// TIA Portal project "S7_1516_LECTOR620_DI" (V15) (continued)
VERSION : 1.2
// The function block use a Profinet/Probibus connection to communicate with a SICK AutoIdent
// device. The FB makes it possible to send and receive sensor data. The Confirmed Messaging 
// protocol (CM-Protocol) is used to receive even long fragmented read results.
// The function block use a Profinet/Probibus connection to communicate with a SICK AutoIdent
// device. The FB makes it possible to send and receive sensor data.
   VAR_INPUT
      HWInputIdent : Hw_Io;   // Hardware identification number of the input module
      HWInputLength : USInt;   // Size of the input module
      HWOutputIdent : Hw_Io;   // Hardware identification number of the output module
      HWOutputLength : USInt;   // Size of the output module
      TOut : Time := T#5s;   // Time out
      Req : Bool;   // A positive edge starts the request
      CommandLength : UInt;   // Byte length of the command / Command length in byte
   END_VAR
   VAR_OUTPUT
      RdDone : Bool;   // Reading result arrived / Positive edge: A reading result sent by the device was received
      RdLength : Int;   // Byte length of the reading result / Length of the reading result in byte
      ReqDone : Bool;   // Requested data available / Indicates whether a CoLa command was sent and an answer was received
      ReqBusy : Bool;   // Request busy / Request processing
      ReqLength : Int;   // Byte length of the requested data / Length of an answer telegram in byte
      Error : Bool;   // Error / Error detected
      Errorcode : DWord;   // Error code / Error code (see documentation)
   END_VAR
   VAR_IN_OUT
      arrCommand : Array[0..499] of Byte;   // Contain the transmitted CoLa command without STX/ETX framing
      arrRecord : Array[0..499] of Byte;   // Contain the received telegram
   END_VAR
   VAR
      bTriggerReq : Bool := false;   // Rising edge detection
      bTriggerReqMem : Bool := false;   // Rising edge detection
      bReadFrag : Bool;   // Fragmentation is needed (Read)
      bWriteFrag : Bool;   // Fragmentation is needed (Write)
      bReqBusyMem : Bool;
      iReadStep : USInt;   // Current step (Read)
      iWriteStep : USInt;   // Current step (Write)
      iReadIndex : UInt;   // Index (Read)
      iWriteIndex : UInt;   // Index (Write)
      iReadHeaderLength : UInt;   // Header length of the CM-Protocol (Read)
      iWriteHeaderLength : UInt;   // Header length of the CM-Protocol (Write)
      iReadFragmentLength : UInt;   // Length of the current fragment (Read)
      iWriteFragmentLength : UInt;   // Length of the current fragment (Write)
      iRecordSize : UInt;   // Length of the record array
      iCommandSize : UInt;   // Length of the command array
      nTempErrorCode : DWord;   // Temporarily error code
      arrInputImage : Array[0..127] of Byte;   // Process data input image
      arrOutputImage : Array[0..127] of Byte;   // Process data output image
      fbTimeout : TON_TIME;   // Instance: Timer on delay (Time out)
   END_VAR
   VAR_TEMP
      iTemp1 : Int;   // Temporarily variable
      iTemp2 : UDInt;   // Temporarily variable
      iTemp3 : UDInt;   // Temporarily variable
   END_VAR
BEGIN
   (*===========================================================================================
   Name:   SICK_CCOMM_PNDP
   Author: SICK AG
   =============================================================================================
   Description: 
   The function block use a Profinet/Probibus connection to communicate with a SICK AutoIdent
   device. The FB makes it possible to send and receive sensor data. The Confirmed Messaging 
   protocol (CM-Protocol) is used to receive even long fragmented read results.

   Send a command:
   The "Req" parameter must be triggered with a rising edge (signal change FALSE to TRUE) in 
   order to carry out the function. For the time during which a valid response has yet to be 
   received from the device, the "ReqBusy" parameter is used to signal  that a response is still 
   pending. The module signals the "ReqDone" = TRUE output parameter when the function has been 
   successfully completed. If data was requested by the device, this data is copied into the 
   Record (arrRecord). The "ReqDone" indicates that new data has been received  for a PLC cycle.
   Only one CoLa-A command request can be send to the same device at one time. 

   Receive a reading result:
   Data sent via trigger command or directly by the device (e.g., direct trigger via a light 
   barrier) is stored in the Record (arrRecord). The "RdDone" output indicates that new data 
   has been received for a PLC cycle. The data sent by the device can be changed or adapted in 
   output format of SOPAS-ET. 

   This AOI supports the folowing SICK devices:
   - Lector6xx
   - RFU6xx
   - CLV6xx 
   - RFH6xx
   =============================================================================================
   Confirmed Messaging Protocol definitions:
   arrInputImage[0]        = Status byte 
   arrInputImage[1]        = Receive counter
   arrInputImage[2]        = Transmit counter back
   arrInputImage[3]        = Command length LSB
   arrInputImage[4]        = Command length MSB
   arrInputImage[5..127]   = Device response (CoLa-A)

   arrOutputImage[0]       = Status byte 
   arrOutputImage[1]       = Receive counter back
   arrOutputImage[2]       = Transmit counter
   arrOutputImage[3]       = Command length LSB
   arrOutputImage[4]       = Command length MSB
   arrOutputImage[5..127]  = Device request (CoLa-A)
   =============================================================================================
   Version history:
   Date       | Version | Created under               | Author  | Remark
   ---------------------------------------------------------------------------------------------
   16/01/2014 | V1.0    | TIA Portal V12 SP1 Update 2 | SICK AG | Initial version
   07/08/2014 | V1.1    | TIA Portal V12 SP1 Update 4 | SICK AG | Replace R_TRIG function 
   22/04/2015 | V1.2    | TIA Portal V12 SP1 Update 4 | SICK AG | Avoid warnings that occur with 
                                                                  TIA V13
   ============================================================================================*)

   (*===================================== INITIALISATION =====================================*)
   #iRecordSize:= 500;   (*Length of the arrRecord array*)
   #iCommandSize:= 500;  (*Length of the arrCommand array*)

   #RdDone:= false;
   #iReadStep:= 0;

   (*Rising edge detection of the request flag*)
   #bTriggerReq:= #Req AND NOT #bTriggerReqMem;
   #bTriggerReqMem:= #Req;

   (*Error detection*)
   IF #nTempErrorCode <>16#0000_0000 THEN
     #ReqDone:= false;
     #ReqBusy:= false;
     #bReqBusyMem:= false;
     #Error:= true;
     #Errorcode:= #nTempErrorCode;
     #nTempErrorCode:= 16#0000_0000;
     #ReqLength:= 0;
     #iWriteStep:= 0;
     RETURN;
   END_IF;

   (*Time out detection*)
   #fbTimeout(IN:=#bReqBusyMem, PT:=#TOut);
   IF #fbTimeout.Q THEN
     #nTempErrorCode:= 16#0000_0001; (*Error: Time out*) 
   END_IF;

   (*Check the hardware ident length of the input module*)
   IF #HWInputLength <8 OR #HWInputLength >128 THEN
     #nTempErrorCode:= 16#0000_0002; (*Error: Incorrect module input length*)
   END_IF;

   (*Check the hardware ident length of the output module*)
   IF #HWOutputLength <8 OR #HWOutputLength >128 THEN
     #nTempErrorCode:= 16#0000_0003; (*Error: Incorrect module output length*)
   END_IF;

   (*Error detected*)
   IF #nTempErrorCode <>16#0000_0000 THEN
     RETURN;
   END_IF;


   (*===================================== COMMUNICATION ======================================*)
   (*Set output data*)
   #iTemp1:= DPWR_DAT(LADDR:= #HWOutputIdent, RECORD:= #arrOutputImage);
   IF #iTemp1 <>0 THEN
     #nTempErrorCode.%W1:= #iTemp1;
     #nTempErrorCode.%W0:= 16#0004; (*Error: Set output data via DPWR_DAT*)
     RETURN;
   END_IF;

   (*Get input data*)
   #iTemp1:= DPRD_DAT(LADDR:= #HWInputIdent, RECORD=> #arrInputImage);
   IF #iTemp1 <>0 THEN
     #nTempErrorCode.%W1:= #iTemp1;
     #nTempErrorCode.%W0:= 16#0005; (*Error: Get input data via DPRD_DAT*)
     RETURN;
   END_IF;

   (*Receive counter ==0 && Receive counter back <>0*)
   IF #arrInputImage[1] =0 AND #arrOutputImage[1] <>0 THEN
     #arrOutputImage[1]:= #arrInputImage[1]; (*Recive counter => Receive counter back*)
     RETURN;
   END_IF;

   (*Transmit counter <> Transmit counter back*)
   IF NOT #bReqBusyMem AND (#arrInputImage[2] <> #arrOutputImage[2]) THEN
     #arrOutputImage[2]:= 0; (*0 => Transmit counter*)
     RETURN;
   END_IF;


   (*============================== HANDLING OF THE RECEIVED DATA =============================*)
   (*New telegram available*)
   IF NOT (#arrInputImage[1] = #arrOutputImage[1]) THEN

     (*Reset error every incoming telegram (Read only mode, e.g. for hand held scanners)*)
     IF #CommandLength <=0 THEN
       #Error:= false;
       #Errorcode:= 16#0000_0000;
     END_IF;

     (*Confirm the receive counter*)
     #arrOutputImage[1]:= #arrInputImage[1];

     (*Get telegram length from the received header*)
     #iReadHeaderLength.%B0:= #arrInputImage[3];
     #iReadHeaderLength.%B1:= #arrInputImage[4];

     (*Check if fragmentation is not active at the moment*)
     IF NOT #bReadFrag THEN
       #iReadIndex:= 0;

       (*Check if fragmentation is needed*)
       IF (#HWInputLength-5) < #iReadHeaderLength THEN
         #bReadFrag:= true;
       END_IF;
     END_IF;

     (*Fragmentation is needed*)
     IF #bReadFrag THEN
       IF (#HWInputLength-5) < #iReadHeaderLength THEN
         #iReadFragmentLength:= #HWInputLength-5;
       ELSE
         #iReadFragmentLength:= #iReadHeaderLength;
       END_IF;

     (*No fragmentation needed*)
     ELSE
       #iReadFragmentLength:= #iReadHeaderLength;
     END_IF;

     (*Copy input data into the output record*)
     IF (#iReadIndex+#iReadFragmentLength) <= #iRecordSize THEN
       MOVE_BLK(IN:= #arrInputImage[5], COUNT:= #iReadFragmentLength, OUT=> #arrRecord[#iReadIndex]);
     END_IF;

     (*Check if all data has been received*)
     IF (#HWInputLength-5) < #iReadHeaderLength THEN
       #iReadIndex:= #iReadIndex+#iReadFragmentLength;

     (*All data has been received*)
     ELSE
       #bReadFrag:= false;
       #iReadStep:= 1;
     END_IF;

     (*Incoming data filter*)
     (* - Check if the receiving telegram os a CoLa answer on a requested 
          comand or a reading result.

         sRA  sWA  sMA  sAN  sAI  sEA  sPX  s{   sSI  sSN  sFA
     sRN  X                                       X    X    X
     sRI  X                                       X    X    X
     sWN       X                                  X    X    X
     sWI       X                                  X    X    X
     sMN            X    X                        X    X    X
     sMI            X         X                   X    X    X
     sEN                           X              X    X    X
     sEI                           X              X    X    X
     sPE                                X         X    X    X
     s{                                      X    X    X    X
     *)
     IF #iReadStep =1 THEN
       (*Filter is only active, while requested data expected*)
       IF #bReqBusyMem THEN
         IF #CommandLength >3 THEN
           (*Get the prefix from the requested command (e.g. 'sRN '*)   
           #iTemp2.%B3:= #arrCommand[0];
           #iTemp2.%B2:= #arrCommand[1];
           #iTemp2.%B1:= #arrCommand[2];
           #iTemp2.%B0:= 16#20;

           (*Get the prefix from the command response (e.g. 'sRA ')*)
           #iTemp3.%B3:= #arrRecord[0];
           #iTemp3.%B2:= #arrRecord[1];
           #iTemp3.%B1:= #arrRecord[2];
           #iTemp3.%B0:= 16#20;
         ELSE
           #iTemp2:= 16#0000_0000;
           #iTemp3:= 16#0000_0000;
         END_IF;

         CASE #iTemp3 OF
         (*'s{  '*)
         16#737B2020:  IF #iTemp2 = 16#737B2020 THEN
                         #iReadStep:= 2; (*Command response*)
                       ELSE
                         #iReadStep:= 3; (*Reading result*)
                       END_IF;

         (*'sRA '*)
         16#73524120:  IF (#iTemp2 = 16#73524E20) OR (#iTemp2 = 16#73524920) THEN
                         #iReadStep:= 2; (*Command response*)
                       ELSE
                         #iReadStep:= 3; (*Reading result*)
                       END_IF;

         (*'sWA '*)
         16#73574120:  IF (#iTemp2 = 16#73574E20) OR (#iTemp2 = 16#73574920) THEN
                         #iReadStep:= 2; (*Command response*)
                       ELSE
                         #iReadStep:= 3; (*Reading result*)
                       END_IF;

         (*'sMA '*)
         16#734D4120:  IF (#iTemp2 = 16#734D4E20) OR (#iTemp2 = 16#734D4920) THEN
                         #iReadStep:= 2; (*Command response*)
                       ELSE
                         #iReadStep:= 3; (*Reading result*)
                       END_IF;

         (*'sAN '*)
         16#73414E20:  IF #iTemp2 = 16#734D4E20 THEN
                         #iReadStep:= 2; (*Command response*)
                       ELSE
                         #iReadStep:= 3; (*Reading result*)
                       END_IF;

         (*'sAI '*)
         16#73414920:  IF #iTemp2 = 16#734D4920 THEN
                         #iReadStep:= 2; (*Command response*)
                       ELSE
                         #iReadStep:= 3; (*Reading result*)
                       END_IF;

         (*'sEA '*)
         16#73454120:  IF (#iTemp2 = 16#73454E20) OR (#iTemp2 = 16#73454920) THEN
                         #iReadStep:= 2; (*Command response*)
                       ELSE
                         #iReadStep:= 3; (*Reading result*)
                       END_IF;

         (*'sPX '*)
         16#73505820:  IF #iTemp2 = 16#73504520 THEN
                         #iReadStep:= 2; (*Command response*)
                       ELSE
                         #iReadStep:= 3; (*Reading result*)
                       END_IF;

         (*'sSI '*)
         16#73534920:  #iReadStep:= 3; (*Reading result*)

         (*'sSN '*)
         16#73534E20:  #iReadStep:= 3; (*Reading result*)

         (*'sFA '*)
         16#73464120:  #iReadStep:= 2; (*Command response*)

         (*Invalid CoLa-A answer*)
         ELSE
           (*Check if a user defined command is used (Request == Response)*)
           FOR #iTemp1:= 0 TO UINT_TO_INT(#CommandLength-1) DO
             IF #arrCommand[#iTemp1] = #arrRecord[#iTemp1] THEN
               #iReadStep:= 2; (*Command response*)
             ELSE
               #iReadStep:= 3; (*Reading result*)
               EXIT;
             END_IF;
           END_FOR;
         END_CASE;

       (*Reading result*)
       ELSE
         #iReadStep:= 3;  (*Reading result*)
       END_IF;
     END_IF;

     (*Incoming telegram is a command response*)
     IF #iReadStep =2 THEN
       IF (#iReadIndex+#iReadFragmentLength) <= #iRecordSize THEN
         #ReqLength:= UDINT_TO_INT(#iReadIndex+#iReadFragmentLength);
         #ReqDone:= true;
         #ReqBusy:= false;
         #bReqBusyMem:= false;
       ELSE
         #nTempErrorCode:= 16#0000_0006; (*Error: Incoming command response > Record size*)
       END_IF;
     END_IF;

     (*Incoming telegram is a reading result*)
     IF #iReadStep =3 THEN
       IF (#iReadIndex+#iReadFragmentLength) <= #iRecordSize THEN
         #RdLength:= UDINT_TO_INT(#iReadIndex+#iReadFragmentLength);
         #RdDone:= true;
       ELSE
         #RdLength:= -1;
         #RdDone:= false;    
       END_IF;
     END_IF;
   END_IF;


   (*=========================== HANDLING OF THE DATA TO BE WRITTEN ===========================*)
   IF #bTriggerReq AND NOT #bReqBusyMem THEN
     #ReqDone:= false;
     #ReqBusy:= true;
     #bReqBusyMem:= true;
     #Error:= false;
     #Errorcode:= 16#0000_0000;
     #iWriteIndex:= 0;

     (*Check command length*)
     IF #CommandLength <=0 THEN
       #nTempErrorCode:= 16#0000_0007; (*Error: Command length <= 0*)
       RETURN;
     ELSIF #CommandLength > #iCommandSize THEN
       #nTempErrorCode:= 16#0000_0008; (*Error: Command length > command array*)
       RETURN;
     END_IF;

     (*Check if the the command telegram must be fragmented*)
     IF (#HWOutputLength-5) < #CommandLength THEN
       #iWriteFragmentLength:= #HWOutputLength-5;
     ELSE
       #iWriteFragmentLength:= #CommandLength;
     END_IF;

     #iWriteHeaderLength:= #CommandLength;
     #iWriteStep:= 1;  
   END_IF;

   (*Write step 1: Command transfer*)
   IF (#iWriteStep =1) AND(#arrInputImage[2] = #arrOutputImage[2]) THEN

     (*Copy command data into the output record*)
     IF((#iWriteIndex+#iWriteFragmentLength) <= #iCommandSize) AND (#iWriteFragmentLength <= (#HWOutputLength-5)) THEN
       MOVE_BLK(IN:= #arrCommand[#iWriteIndex], COUNT:= #iWriteFragmentLength, OUT=> #arrOutputImage[5]);
       (*Increment transmit counter*)
       IF #arrOutputImage[2] = 16#FF THEN
         #arrOutputImage[2]:= 16#01; (*Counter overflow, zero is skipped*)
       ELSE
         #arrOutputImage[2]:= #arrOutputImage[2]+1;
       END_IF;

       (*Set command/fragment length*)
       #arrOutputImage[3]:= #iWriteHeaderLength.%B0;
       #arrOutputImage[4]:= #iWriteHeaderLength.%B1;

       (*Next step*)
       #iWriteStep:= 2;
     ELSE
       #nTempErrorCode:= 16#0000_0009; (*Error: Fragmentation error*)
     END_IF;
       RETURN;
   END_IF;

   (*Write step 2: Fragmentation handling*)
   IF #iWriteStep =2 THEN

     (*Fragmentation is needed*)
     IF (#HWOutputLength-5) < #iWriteHeaderLength THEN
       #bWriteFrag:= true;

       (*Next index*)
       #iWriteIndex:= #iWriteIndex+#iWriteFragmentLength;

       (*Set next header length*)
       #iWriteHeaderLength:= #iWriteHeaderLength-#iWriteFragmentLength;

       (*Set next fragment length*)
       IF (#HWOutputLength-5) < #iWriteHeaderLength THEN
         #iWriteFragmentLength:= #HWOutputLength-5;
       ELSE
         #iWriteFragmentLength:= #iWriteHeaderLength;
       END_IF;

     (*Fragmentation is not needed*)
     ELSE
       #bWriteFrag:= false;
     END_IF;

     (*Next step*)
     #iWriteStep:= 3;
   END_IF;

   (*Write step 3: Check if the transmission of the command/fragment is done*)
   IF #iWriteStep =3 THEN

     (*Transmit counter back == Transmit counter*)
     IF #arrInputImage[2] = #arrOutputImage[2] THEN
       IF #bWriteFrag THEN
         #iWriteStep:= 1;
       ELSE
         #iWriteStep:= 0;
       END_IF;
     END_IF;
   END_IF;
END_FUNCTION_BLOCK

FUNCTION "SICK_GetValue" : Void   // FC10, SCL
TITLE = Get value
{ S7_Optimized_Access := 'TRUE' }
AUTHOR : SICKAG
FAMILY : Ident
VERSION : 1.0
// This function is needs to get a value out of a SICK CoLa command.
   VAR_INPUT
      iTelegramLength : UInt;   // Length of the source telegram
      iValueLength : USInt;   // ASCII length of the value [1..8] = Fix length | [0]= Variable
      arrData : Array[0..499] of Byte;   // Data record (contains the whole CoLa telegram)
   END_VAR
   VAR_OUTPUT
      nValue : DWord;   // Read value
      nErrorCode : Word;   // Error code
   END_VAR
   VAR_IN_OUT
      iPosition : UInt;   // Position offset of the value before and after (starting from 0)
   END_VAR
   VAR_TEMP
      iLoop : Int;   // Temporarily variable
      iSegmentLength : UInt;   // Length of the segement
      nTemp : DWord;   // Temporarily variable
   END_VAR
BEGIN
   (*===========================================================================================
   Name:   SICK_GetValue
   Author: SICK AG
   =============================================================================================
   Description: 
   This function is for internal use only. The function gets the selected Hex-value string out 
   of the CoLa-Telegram and convert it into a hexadecimal number. 

   =============================================================================================
   Error codes:
   16#0000 = No error
   16#0001 = Invaild telegram length   
   16#0002 = Invalid position index 
   16#0003 = Invalid value length
   16#0004 = Invalid segment length 
   16#0005 = ASCII character is not in a hexadecimal format             

   =============================================================================================
   Version history:
   Date       | Version | created under               | Author  | Remark
   ---------------------------------------------------------------------------------------------
   30/01/2014 | V1.0    | TIA Portal V12 SP1 Update 2 | SICK AG | Initial version
   ============================================================================================*)

   (*===================================== INITIALISATION =====================================*)
   #iSegmentLength:= 0;
   #nValue:= 16#0000_0000;
   #nErrorCode:= 16#0000;

   (*======================================= READ VALUE =======================================*)
   (*Check telegram length*)
   IF #iTelegramLength <=0 OR #iTelegramLength > 500 THEN
     #nErrorCode:= 16#0001; (*Error: Invaild telegram length*)
     RETURN;
   END_IF;

   (*Check current position of the value*)
   IF #iPosition > (#iTelegramLength-1) THEN
     #nErrorCode:= 16#0002; (*Error: Invalid position index*)
     RETURN;
   END_IF;

   (*Check value length*)
   IF #iValueLength >8 THEN
     #nErrorCode:= 16#0003; (*Error: Invalid value length*)
     RETURN;
   END_IF;

   (*Get a value with a variable length (ends with a ' ' or [ETX]*)
   IF #iValueLength = 0 THEN
     FOR #iLoop:= UINT_TO_INT(#iPosition) TO UINT_TO_INT(#iTelegramLength-1) DO
       (*Check if a blank or a [ETX] is detected*)
       IF (#arrData[#iLoop] =' ') OR (#arrData[#iLoop] ='$03') THEN
         EXIT;
       END_IF;

       (*Length of the current value segement*)
       #iSegmentLength:= #iSegmentLength+1;
     END_FOR;

   (*Get a value with a fixed character length [1..8]*)
   ELSE
     #iSegmentLength:= #iValueLength;
   END_IF;

   (*Check if the segment length is valid*)
   IF (#iSegmentLength >8) OR (#iSegmentLength =0) THEN
     #nErrorCode:= 16#0004; (*Error: Invalid segment length*)
     RETURN;
   END_IF;

   (*Convert ASCII string into a hexadecimal number*)
   FOR #iLoop:= UINT_TO_INT(#iPosition) TO UINT_TO_INT(#iPosition+#iSegmentLength-1) DO
     (*ACSII value = [0..9]*)
     IF #arrData[#iLoop] >='0' AND #arrData[#iLoop] <='9' THEN
       #nTemp:= #arrData[#iLoop]-48;
     (*ASCII value = [A..F]*) 
     ELSIF #arrData[#iLoop] >='A' AND #arrData[#iLoop] <='F' THEN
       #nTemp:= #arrData[#iLoop]-55;
     (*ASCII value = [a..f]*)
     ELSIF #arrData[#iLoop] >='a' AND #arrData[#iLoop] <='f' THEN
       #nTemp:= #arrData[#iLoop]-87;    
     ELSE
       #nErrorCode:= 16#0005; (*Error: ASCII character is not in a hexadecimal format *)
       RETURN;
     END_IF;

     (*Create hexadecimal number*)
     #nValue:= SHL(IN:= #nValue, N:= 4);
     #nValue:= #nValue+#nTemp;
   END_FOR;

   (*Set the position of the next element in the telegram*)
   IF #iValueLength = 0 THEN
     #iPosition:= #iPosition+#iSegmentLength+1; (*With blank character*)
   ELSE
     #iPosition:= #iPosition+#iSegmentLength; (*Without blank character*)
   END_IF;
END_FUNCTION

FUNCTION "SICK_SetValue" : Void   // FC11, SCL
TITLE = Set value
{ S7_Optimized_Access := 'TRUE' }
AUTHOR : SICKAG
FAMILY : Ident
VERSION : 1.1
// This function is needs to set a value to a SICK CoLa command.
   VAR_INPUT
      bAddBlank : Bool;   // Add blank after value
      nValue : DWord;   // Value that should be written
   END_VAR
   VAR_OUTPUT
      arrData : Array[0..499] of Byte;   // Destination telegram
      nErrorCode : Word;   // Error code
   END_VAR
   VAR_IN_OUT
      iPosition : UInt;   // Position offset of the value before and after (starting from 0)
   END_VAR
   VAR_TEMP
      iValueLength : USInt;   // Byte length of the value that shuld be written
      nReturnValue : Word;   // Return value of the convert function
      sValue : String[8];   // Converted value
      nTempValue : DWord;   // Temporarily variable
      iTemp : UInt;   // Temporarily variable
   END_VAR
BEGIN
   (*===========================================================================================
   Name:   SICK_SetValue
   Author: SICK AG
   =============================================================================================
   Description: 
   This function is for internal use only.
   The function converts a hexadecimal value into a hexadecimal string and add it 
   automatically to the command array.     

   =============================================================================================
   Error codes:
   16#0000 = No error
   16#0001 = Invalid position index   
   16#8xxx = Conversion error (HTA-Function) see help system for more information

   =============================================================================================
   Version history:
   Date       | Version | created under               | Author  | Remark
   ---------------------------------------------------------------------------------------------
   30/01/2014 | V1.0    | TIA Portal V12 SP1 Update 2 | SICK AG | Initial version
   22/04/2014 | V1.1    | TIA Portal V12 SP1 Update 4 | SICK AG | Avoid warnings that occur with 
                                                                  TIA V13
   ============================================================================================*)

   (*===================================== INITIALISATION =====================================*)
   #iValueLength:= 0;
   #nErrorCode:= 16#0000;

   (*======================================= WRITE VALUE ======================================*)
   (*Check current position of the value*)
   IF #iPosition > 499 THEN 
     #nErrorCode:= 16#0001; (*Error: Invalid position index*)
     RETURN;
   END_IF;



   (*Get byte length of the value that should be written*)
   IF #nValue <= 16#FF THEN
     #nTempValue:= SHL(IN:= #nValue, N:=24);
     #iValueLength:= 1;
   ELSIF #nValue <= 16#FFFF THEN
     #nTempValue:= SHL(IN:= #nValue, N:=16);
     #iValueLength:= 2;
   ELSIF #nValue <= 16#00FF_FFFF THEN
     #nTempValue:= SHL(IN:= #nValue, N:=8);
     #iValueLength:= 3;
   ELSIF #nValue <= 16#FFFF_FFFF THEN
     #nTempValue:= #nValue;
     #iValueLength:= 4;
   END_IF;

   (*Convert hexadecimal number into a ASCII string*)
   #nReturnValue:= HTA(IN:= #nTempValue, N:= #iValueLength, OUT=>#sValue);
   IF #nReturnValue <> 16#0000 THEN
     #nErrorCode:= #nReturnValue; (*Error: Conversion error (HTA-Function)*)
     RETURN;
   END_IF;

   (*Add the string value to the destination telegram*)
   #arrData[#iPosition]:= 0; // Avoid warnings under TIA V13
   Strg_TO_Chars(Strg:=#sValue, pChars:= #iPosition, Cnt=> #iTemp, Chars:= #arrData);

   (*Add blank to the destination telegram and calculate the position of the next element*)
   IF #bAddBlank THEN
     #arrData[#iPosition+#iTemp]:= ' ';
     #iPosition:= #iPosition+#iTemp+1;

   (*Calculate the position of the next element*)
   ELSE
     #iPosition:= #iPosition+#iTemp;
   END_IF;
END_FUNCTION

(* ===== HMI "HMI_RT_1" =====
system functions are stored by id; their names below are inferred from use
connection "HMI_Connection_1": ETHERNET, S7_1500_OMS

HMI tags "Default tag table"
   "No_of_counts_in" : Byte = PLC No_of_counts_in AT %IB57, 1 s
   "iCounter_Tag_kopija" : Int = PLC iCounter_Tag_kopija AT %QW12, 1 s
   "Sensor_ok_blinking" : Byte = PLC Data_block_1.Sensor_ok_blink AT %DB1.DBB7, 500 ms

HMI tags "Lector620"
   "PocasniPrebranaKoda" : String[254] = PLC Data_block_1.ShranjenaPrebranaKoda AT %DB1.DBX54.0, 500 ms
   "Rocno_Prozenje" : Bool = PLC Data_block_1.TestBitStefanRequest AT %DB1.DBX44.0, 1 s

Template "Template" 800x480
   GraphicView "Template_Graphic view_1" at 0,0 size 466x201; Picture "Image_0246DFF1_1EB2_3537_41B2_099D4BE026E4 (1)"
   Clock "Template_Clock_1" at 514,13 size 219x137
   DateTimeField "Template_Date/time field_1" at 508,173 size 241x32

screen "Lector_HMI_Start" 800x480, template "Template"
   IOField "I/O field_1" at 49,406 size 706x61; FormatPattern ???????????????????????????????????????????????????????????????????????????????????????????????????????????????????????????????????????????????????????????????????????????????????????????????????????????????????????????????????????????????????????????????
      ProcessValue <- "PocasniPrebranaKoda"
   Circle "Circle_1" at 498,338 size 43x43
      Appearance <- "Sensor_ok_blinking"
   Button "Button_1" at 644,335 size 96x32; TextOff 'Exit RT'
      on Click: StopRuntime(0)
   Button "Button_2" at 295,243 size 157x75; TextOff 'Rocno Prozenje'
      on Press: function_b14e0dd5("Rocno_Prozenje", 0)
   TextField "Text Field_6" at 231,338 size 240x43; Text 'Nr. / No. / Senzor Aktiven'
*)

(* ===== HMI "HMI_RT_2" =====
system functions are stored by id; their names below are inferred from use
connection "HMI_Connection_2": ETHERNET, S7_1500_OMS

HMI tags "Default tag table"
   "SICK_IN_1" : Bool = PLC SICK_IN_1 AT %Q0.0, 1 s

HMI tags "Lector_PC_Tags"
   "ID" : Array [0..5] of Int, internal   // ID stevilke
   "Serijska_Stevilka_0" : WString[255], internal   // Pozor da length bode nastavljen koliko je potrebno
   "Serijska_Stevilka_1" : WString[255], internal
   "Serijska_Stevilka_2" : WString[255], internal
   "Serijska_Stevilka_3" : WString[255], internal
   "Serijska_Stevilka_4" : WString[255], internal
   "Serijska_Stevilka_5" : WString[255], internal
   "Stevilo_Branja" : Array [0..5] of Int, internal   // Stevilo branja iste kode
   "Cas_Poslednjega_Branja" : Array [0..5] of DateTime, internal   // Datum in cas poslednjega branja kode
   "szDatabase" : WString[30], internal   // Ime baze podatkov
   "szTableName" : WString[30], internal   // Ime tabele v bazi podatkov
   "Count_Number" : LInt = PLC Data_block_1.No_of_counts AT %DB1.DBX8.0, 100 ms
      on ChangeValue: SetTag("Novi_Artikel_Koda_Artikla_Temp", "PrebranaKoda"); "Sprejem_Serijske_Stevilke_v_SQL"('Database_ArchiveMessage')
   "nTab" : Int, internal   // Sledi scrollanje tabela
   "PrebranaKoda" : String[254] = PLC Data_block_1.ShranjenaPrebranaKoda AT %DB1.DBX54.0, 100 ms
   "PocasniPrebranaKoda" : String[254] = PLC Data_block_1.ShranjenaPrebranaKoda AT %DB1.DBX54.0, 1 s
   "PrebranaKoda_Cas" : Date_And_Time = PLC Data_block_1.ShranjenaPrebranaKoda_Cas AT %DB1.DBX46.0, 100 ms
   "temp" : WString[10] AT %DB1.DBX0.0
   "Ime_Artikla_0" : WString[255], internal   // Pozor da length bode nastavljen koliko je potrebno
   "Ime_Artikla_1" : WString[255], internal
   "Ime_Artikla_2" : WString[255], internal
   "Ime_Artikla_3" : WString[255], internal
   "Ime_Artikla_4" : WString[255], internal
   "Ime_Artikla_5" : WString[255], internal
   "Stanje_0" : WString[255], internal
   "Stanje_1" : WString[255], internal
   "Stanje_2" : WString[255], internal
   "Stanje_3" : WString[255], internal
   "Stanje_4" : WString[255], internal
   "Stanje_5" : WString[255], internal
   "Ime_Artikla_temp" : WString[255], internal
   "Stanje_temp" : WString[255], internal
   "tempID_Tag" : Array [0..5] of Int, internal
   "Iskanje_ID" : Int, internal
   "Iskanje_Instanci" : WString[255], internal
   "ID_Instance" : Array [0..5] of Int, internal
   "Prebrana_Koda_FLAG" : Bool = PLC Data_block_1.Prebrana_Koda_FLAG AT %DB1.DBX318.0   // Pri Value Change Event-u aktivira scriptu za sprejem
   "Stanje_Update_Select" : Int, internal
   "Rocno_Prozenje" : Bool = PLC Data_block_1.TestBitStefanRequest AT %DB1.DBX44.0, 500 ms
   "Startup_Setup" : Bool AT %DB1.DBX0.0

HMI tags "PopUp_tags"
   "Naredi_Novi_Artikel_DA" : Bool, internal
   "Nova_Serijska_Stevilka_Prebrana_ALARM" : Int, internal
   "Popup_Naredi_Novi_Artikel" : Bool, internal   // Spremeni ga alarm za branje nove kode
      on ChangeValue: function_f294b399("Naredi_Nov_Artikel", 0, 0, 1280, 1024, -1, -1, 1)
   "Novi_Artikel_Ime_Artikla_Temp" : WString[255], internal
   "Novi_Artikel_ID_Artikla_Temp" : Int, internal
   "Novi_Artikel_Stanje_Artikla_Temp" : WString[255], internal
   "Novi_Artikel_Koda_Artikla_Temp" : WString[255], internal

discrete alarms
   1: 'Nova serijska stevilka prebrana, katera ne obstaja v sistemu', class Warnings, trigger "Nova_Serijska_Stevilka_Prebrana_ALARM" bit 0
      on Coming: SetTag("Popup_Naredi_Novi_Artikel", 1)

screen "Lector_zacetek" 1280x1024, template "Template_LectorStart"
   on GenerateScreen: function_a9b64e44("Nova_Serijska_Stevilka_Prebrana_ALARM", 0); ResetBit("Prebrana_Koda_FLAG"); ResetBit("Popup_Naredi_Novi_Artikel"); "RT_Startup_Setup"()
   Button "Button_1" at 12,935 size 96x72; TextOff 'IZHOD'
      on Press: StopRuntime(0)
   Button "Button_2" at 540,380 size 200x87; TextOff 'SQL Tabele'
      on Click: ActivateScreen("Lector_Branje_Tabela", 0)
   IOField "I/O field_1" at 11,543 size 1251x61; FormatPattern ????????????????????????????????????????????????????????????????????????????????????????????????????????????????????????????????????????????????????????????????????????????????????????????????????????
      ProcessValue <- "PocasniPrebranaKoda"
   Button "FB_Information_Round" at 1175,935 size 72x72; TextOff 'Text'; PictureOn "FB_Information_Round_Pressed_256c"; PictureOff "FB_Information_Round_Released_256c"

Template "Template_Support" 1280x1024
   TextField "_Vorlage_Textfeld_1" at 25,45 size 37x332; Text 'Industry Online Support'

Template "Template_LectorStart" 1280x1024
   GraphicView "Template_Graphic view_1" at 316,0 size 633x307; Picture "Image_0246DFF1_1EB2_3537_41B2_099D4BE026E4 (1)"
   Clock "Template_Clock_1" at 1013,33 size 232x220

screen "Lector_Branje_Tabela" 1280x1024, template "Template_LectorStart"
   on GenerateScreen: "Branje_Artiklov"('Database_ArchiveMessage')
   IOField "IO Field" at 279,519 size 214x43; FormatPattern ???????????????????????????????????????????????????????????????????????????????????????????????????????????????????????????????????????????????????????????????????????????????????????????????????????????????????????????????????????????????????????????????
      ProcessValue <- "Ime_Artikla_0"
   IOField "IO Field_0" at 782,516 size 161x43; FormatPattern 9999
      ProcessValue <- "[0]"
   IOField "IO Field_3" at 979,519 size 279x43; FormatPattern 9999
      ProcessValue <- "[0]"
   IOField "IO Field_7" at 26,517 size 219x43; FormatPattern 999
      ProcessValue <- "[0]"
   IOField "IO Field_8" at 279,577 size 214x43; FormatPattern ???????????????????????????????????????????????????????????????????????????????????????????????????????????????????????????????????????????????????????????????????????????????????????????????????????????????????????????????????????????????????????????????
      ProcessValue <- "Ime_Artikla_1"
   IOField "IO Field_10" at 782,574 size 161x43; FormatPattern 9999
      ProcessValue <- "[1]"
   IOField "IO Field_11" at 979,577 size 279x43; FormatPattern 9999
      ProcessValue <- "[1]"
   IOField "IO Field_12" at 26,575 size 219x43; FormatPattern 999
      ProcessValue <- "[1]"
   IOField "IO Field_13" at 279,636 size 214x43; FormatPattern ???????????????????????????????????????????????????????????????????????????????????????????????????????????????????????????????????????????????????????????????????????????????????????????????????????????????????????????????????????????????????????????????
      ProcessValue <- "Ime_Artikla_2"
   IOField "IO Field_14" at 782,633 size 161x43; FormatPattern 9999
      ProcessValue <- "[2]"
   IOField "IO Field_15" at 979,636 size 279x43; FormatPattern 9999
      ProcessValue <- "[2]"
   IOField "IO Field_16" at 26,634 size 219x43; FormatPattern 999
      ProcessValue <- "[2]"
   Button "Button_2" at 1174,313 size 84x70; TextOff 'Text'; PictureOff "Up_Arrow_4"
      on Press: function_b9b71300("nTab", 1); "Scrolling_Up_Down_Artikli"('Database_ArchiveMessage')
   Button "Button" at 1174,935 size 84x70; TextOff 'Text'; PictureOff "Down_Arrow_4"
      on Press: function_dd21b452("nTab", 1); "Scrolling_Up_Down_Artikli"('Database_ArchiveMessage')
   TextField "Text Field_12" at 26,447 size 220x43; Text 'Nr. / No. / ID'
   Button "Button_1" at 32,963 size 143x43; TextOff '<< / Glavni Meni'
      on Press: ActivateScreen("Lector_zacetek", 0)
   IOField "IO Field_9" at 279,695 size 214x43; FormatPattern ???????????????????????????????????????????????????????????????????????????????????????????????????????????????????????????????????????????????????????????????????????????????????????????????????????????????????????????????????????????????????????????????
      ProcessValue <- "Ime_Artikla_3"
   IOField "IO Field_17" at 782,692 size 161x43; FormatPattern 9999
      ProcessValue <- "[3]"
   IOField "IO Field_18" at 979,695 size 279x43; FormatPattern 9999
      ProcessValue <- "[3]"
   IOField "IO Field_19" at 26,693 size 219x43; FormatPattern 999
      ProcessValue <- "[3]"
   IOField "IO Field_20" at 279,753 size 214x43; FormatPattern ???????????????????????????????????????????????????????????????????????????????????????????????????????????????????????????????????????????????????????????????????????????????????????????????????????????????????????????????????????????????????????????????
      ProcessValue <- "Ime_Artikla_4"
   IOField "IO Field_21" at 782,750 size 161x43; FormatPattern 9999
      ProcessValue <- "[4]"
   IOField "IO Field_22" at 979,753 size 279x43; FormatPattern FFFF
      ProcessValue <- "[4]"
   IOField "IO Field_23" at 26,751 size 219x43; FormatPattern 999
      ProcessValue <- "[4]"
   IOField "IO Field_24" at 279,812 size 214x43; FormatPattern ???????????????????????????????????????????????????????????????????????????????????????????????????????????????????????????????????????????????????????????????????????????????????????????????????????????????????????????????????????????????????????????????
      ProcessValue <- "Ime_Artikla_5"
   IOField "IO Field_25" at 782,809 size 161x43; FormatPattern 9999
      ProcessValue <- "[5]"
   IOField "IO Field_26" at 979,812 size 279x43; FormatPattern 9999
      ProcessValue <- "[5]"
   IOField "IO Field_27" at 26,810 size 219x43; FormatPattern 999
      ProcessValue <- "[5]"
   TextField "Text Field_2" at 279,447 size 214x43; Text 'Nr. / No. / Ime Artikla'
   TextField "Text Field_3" at 781,447 size 161x43; Text 'Nr. / No. / Stevilo Branj'
   TextField "Text Field_4" at 979,447 size 279x43; Text 'Nr. / No. / Cas Zadnjega Branja'
   Button "Button_4" at 333,311 size 279x103; TextOff 'Datensatz auslesen / Read data record / Pregled Prebranih Artiklov'
      on Press: ActivateScreen("Lector_Pregled_Prebranih_Artiklov", 0)
   Button "Button_3" at 1009,311 size 109x90; TextOff 'Random'
      on Press: function_b3f726e6("Nova_Serijska_Stevilka_Prebrana_ALARM", 0)
   IOField "IO Field_4" at 518,518 size 244x43; FormatPattern ???????????????????????????????????????????????????????????????????????????????????????????????????????????????????????????????????????????????????????????????????????????????????????????????????????????????????????????????????????????????????????????????
      ProcessValue <- "Serijska_Stevilka_0"
   IOField "IO Field_5" at 518,576 size 244x43; FormatPattern ???????????????????????????????????????????????????????????????????????????????????????????????????????????????????????????????????????????????????????????????????????????????????????????????????????????????????????????????????????????????????????????????
      ProcessValue <- "Serijska_Stevilka_1"
   IOField "IO Field_6" at 518,635 size 244x43; FormatPattern ???????????????????????????????????????????????????????????????????????????????????????????????????????????????????????????????????????????????????????????????????????????????????????????????????????????????????????????????????????????????????????????????
      ProcessValue <- "Serijska_Stevilka_2"
   IOField "IO Field_28" at 518,694 size 244x43; FormatPattern ???????????????????????????????????????????????????????????????????????????????????????????????????????????????????????????????????????????????????????????????????????????????????????????????????????????????????????????????????????????????????????????????
      ProcessValue <- "Serijska_Stevilka_3"
   IOField "IO Field_29" at 518,752 size 244x43; FormatPattern ???????????????????????????????????????????????????????????????????????????????????????????????????????????????????????????????????????????????????????????????????????????????????????????????????????????????????????????????????????????????????????????????
      ProcessValue <- "Serijska_Stevilka_4"
   IOField "IO Field_30" at 518,811 size 244x43; FormatPattern ???????????????????????????????????????????????????????????????????????????????????????????????????????????????????????????????????????????????????????????????????????????????????????????????????????????????????????????????????????????????????????????????
      ProcessValue <- "Serijska_Stevilka_5"
   TextField "Text Field_5" at 518,446 size 244x43; Text 'Nr. / No. / Serijska Stevilka'
   AlarmView "Alarm view_1" at 354,872 size 624x140
   Button "Button_5" at 32,311 size 279x103; TextOff 'Datensatz auslesen / Read data record / Osvezi'
      on Press: "Branje_Artiklov"('Database_ArchiveMessage')
   Button "Button_6" at 636,310 size 279x103; TextOff 'Datensatz auslesen / Read data record / Napredne Funkcije'
      on Click: ActivateScreen("Lector_Napredne_Funkcije", 0)

PopupScreen "Naredi_Nov_Artikel" 600x600
   TextField "Text field_1" at 29,47 size 551x66; Text 'Nova koda je prebrana, katera ni v sistemu. Ali bi zeleli narediti novi artikel za to kodo?'
   Button "Button_1" at 29,223 size 155x89; TextOff 'DA'
      on Click: ActivateScreen("Lector_vnos_novega_artikla", 0); ResetBit("Popup_Naredi_Novi_Artikel")
   Button "Button_2" at 425,223 size 155x89; TextOff 'NE'
      on Click: ResetBit("Prebrana_Koda_FLAG"); function_a9b64e44("Nova_Serijska_Stevilka_Prebrana_ALARM", 0); ResetBit("Popup_Naredi_Novi_Artikel")

screen "Lector_Pregled_Prebranih_Artiklov" 1280x1024
   on GenerateScreen: "Branje_Instanci_Artiklov"('Database_ArchiveMessage')
   IOField "IO Field_0" at 382,517 size 161x43; FormatPattern ????????????????????????????????????????????????????????????????????????????????
      ProcessValue <- "Stanje_0"
      on OnFinishInput: SetTag("Stanje_Update_Select", 0); "Update_Stanja"('Database_ArchiveMessage')
   IOField "IO Field_3" at 559,519 size 279x43; FormatPattern 9999
      ProcessValue <- "[0]"
   IOField "IO Field_7" at 26,517 size 161x43; FormatPattern 999
      ProcessValue <- "[0]"
   IOField "IO Field_10" at 382,575 size 161x43; FormatPattern ????????????????????????????????????????????????????????????????????????????????
      ProcessValue <- "Stanje_1"
      on OnFinishInput: SetTag("Stanje_Update_Select", 1); "Update_Stanja"('Database_ArchiveMessage')
   IOField "IO Field_11" at 559,577 size 279x43; FormatPattern 9999
      ProcessValue <- "[1]"
   IOField "IO Field_12" at 26,575 size 161x43; FormatPattern 999
      ProcessValue <- "[1]"
   IOField "IO Field_14" at 382,634 size 161x43; FormatPattern ????????????????????????????????????????????????????????????????????????????????
      ProcessValue <- "Stanje_2"
      on OnFinishInput: SetTag("Stanje_Update_Select", 2); "Update_Stanja"('Database_ArchiveMessage')
   IOField "IO Field_15" at 559,636 size 279x43; FormatPattern 9999
      ProcessValue <- "[2]"
   IOField "IO Field_16" at 26,634 size 161x43; FormatPattern 999
      ProcessValue <- "[2]"
   Button "Button_2" at 901,364 size 84x70; TextOff 'Text'; PictureOff "Up_Arrow_4"
      on Press: function_b9b71300("nTab", 1); "Scrolling_Up_Down_Instanci"('Database_ArchiveMessage')
   TextField "Text Field_12" at 26,447 size 162x43; Text 'Nr. / No. / ID Artikla'
   IOField "IO Field_17" at 382,693 size 161x43; FormatPattern ????????????????????????????????????????????????????????????????????????????????
      ProcessValue <- "Stanje_3"
      on OnFinishInput: SetTag("Stanje_Update_Select", 3); "Update_Stanja"('Database_ArchiveMessage')
   IOField "IO Field_18" at 559,695 size 279x43; FormatPattern 9999
      ProcessValue <- "[3]"
   IOField "IO Field_19" at 26,693 size 161x43; FormatPattern 999
      ProcessValue <- "[3]"
   IOField "IO Field_21" at 382,751 size 161x43; FormatPattern ????????????????????????????????????????????????????????????????????????????????
      ProcessValue <- "Stanje_4"
      on OnFinishInput: SetTag("Stanje_Update_Select", 4); "Update_Stanja"('Database_ArchiveMessage')
   IOField "IO Field_22" at 559,753 size 279x43; FormatPattern FFFF
      ProcessValue <- "[4]"
   IOField "IO Field_23" at 26,751 size 161x43; FormatPattern 999
      ProcessValue <- "[4]"
   IOField "IO Field_25" at 382,810 size 161x43; FormatPattern ????????????????????????????????????????????????????????????????????????????????
      ProcessValue <- "Stanje_5"
      on OnFinishInput: SetTag("Stanje_Update_Select", 5); "Update_Stanja"('Database_ArchiveMessage')
   IOField "IO Field_26" at 559,812 size 279x43; FormatPattern 9999
      ProcessValue <- "[5]"
   IOField "IO Field_27" at 26,810 size 161x43; FormatPattern 999
      ProcessValue <- "[5]"
   TextField "Text Field_3" at 381,448 size 161x43; Text 'Nr. / No. / Stanje'
   TextField "Text Field_4" at 559,447 size 279x43; Text 'Nr. / No. / Cas Zadnjega Branja'
   DateTimeField "Date/time field_1" at 227,320 size 336x43
   Button "Button" at 836,868 size 84x70; TextOff 'Text'; PictureOff "Down_Arrow_4"
      on Press: function_dd21b452("nTab", 1); "Scrolling_Up_Down_Instanci"('Database_ArchiveMessage')
   IOField "IO Field_4" at 201,517 size 161x43; FormatPattern 999
      ProcessValue <- "[0]"
   IOField "IO Field_5" at 201,575 size 161x43; FormatPattern 999
      ProcessValue <- "[1]"
   IOField "IO Field_6" at 201,634 size 161x43; FormatPattern 999
      ProcessValue <- "[2]"
   TextField "Text Field_2" at 201,447 size 162x43; Text 'Nr. / No. / ID Instance'
   IOField "IO Field_8" at 201,693 size 161x43; FormatPattern 999
      ProcessValue <- "[3]"
   IOField "IO Field_9" at 201,751 size 161x43; FormatPattern 999
      ProcessValue <- "[4]"
   IOField "IO Field_13" at 201,810 size 161x43; FormatPattern 999
      ProcessValue <- "[5]"
   Button "Button_1" at 32,963 size 143x43; TextOff '<<'
      on Press: ActivateScreen("Lector_Branje_Tabela", 0)
   IOField "IO Field_1" at 289,101 size 214x43; FormatPattern ????????????????????????????????????????????????????????????????????????????????????????????????????????????????????????????????????????????????????????????????????????????????????????????????????????????????????????????????????????????????????????????????
      ProcessValue <- "Iskanje_Instanci"
      on OnFinishInput: "Iskanje_po_imenu_artikla"('Database_ArchiveMessage')
   IOField "IO Field_2" at 291,159 size 214x43; FormatPattern 999
      on OnFinishInput: "Iskanje_po_ID"('Database_ArchiveMessage')
      ProcessValue <- "Iskanje_ID"
   TextField "Text Field_1" at 31,159 size 214x43; Text 'Nr. / No. / ID Artikla'
   TextField "Text Field_6" at 31,101 size 214x43; Text 'Nr. / No. / Ime Artikla'
   TextField "Text field_7" at 175,27 size 182x34; Text 'Nacini iskanja'
   Button "Button_3" at 227,963 size 143x43; TextOff '<< / Glavni Meni'
      on Press: ActivateScreen("Lector_zacetek", 0)
   AlarmView "Alarm view_1" at 611,27 size 612x217
   Button "Button_4" at 1011,447 size 260x127; TextOff 'Razvrsti po casu branja'
      on Click: "Branje_Instanci_Artiklov"('Database_ArchiveMessage')

screen "Lector_vnos_novega_artikla" 1280x1024, template "Template_LectorStart"
   on GenerateScreen: SetTag("Novi_Artikel_Ime_Artikla_Temp", 0); SetTag("Novi_Artikel_ID_Artikla_Temp", 0)
   IOField "IO Field_1" at 346,498 size 240x43; FormatPattern ????????????????????????????????????????????????????????????????????????????????????????????????????????????????????????????????????????????????????????????????????????????????????????????????????????????????????????????????????????????????????????????????
      ProcessValue <- "Novi_Artikel_Ime_Artikla_Temp"
   TextField "Text Field_6" at 88,498 size 240x43; Text 'Nr. / No. / Ime Artikla'
   IOField "IO Field_3" at 347,578 size 240x43; FormatPattern 99999
      ProcessValue <- "Novi_Artikel_ID_Artikla_Temp"
   TextField "Text Field_3" at 89,578 size 240x43; Text 'Nr. / No. / Dodeljen ID'
   TextField "Text field_7" at 161,378 size 290x40; Text 'Ustvari novi artikel'
   IOField "IO Field_4" at 401,664 size 834x43; FormatPattern ????????????????????????????????????????????????????????????????????????????????????????????????????????????????????????????????????????????????????????????????????????????????????????????????????????????????????????????????????????????????????????????????
      on OnFinishInput: "Iskanje_po_imenu_artikla"('Database_ArchiveMessage')
      ProcessValue <- "Novi_Artikel_Koda_Artikla_Temp"
   TextField "Text Field_2" at 66,664 size 317x43; Text 'Nr. / No. / Serijska Koda Novega Artikla'
   TextField "Text field_4" at 119,710 size 225x22; Text '(Koda se ne more spremeniti)'
   Button "Button_1" at 636,437 size 302x141; TextOff 'Ustvari artikel na osnovi vnesenih podatkov'
      on Click: "Sprejem_Serijske_Stevilke_v_SQL_Nova_Stevilka"('Database_ArchiveMessage')
   Button "Button_2" at 32,963 size 143x43; TextOff '<< / Nazaj'
      on Press: ResetBit("Prebrana_Koda_FLAG"); function_a9b64e44("Nova_Serijska_Stevilka_Prebrana_ALARM", 0); ResetBit("Popup_Naredi_Novi_Artikel"); SetTag("Novi_Artikel_Ime_Artikla_Temp", '""'); SetTag("Novi_Artikel_Stanje_Artikla_Temp", '""'); ActivateScreen("Lector_zacetek", 0)
   AlarmView "Alarm view_1" at 544,707 size 635x300

screen "Lector_Napredne_Funkcije" 1280x1024, template "Template_LectorStart"
   on GenerateScreen: function_f23ef4c9()
   on ClearScreen: function_f23ef4c9()
   TextField "Text field_1" at 497,342 size 271x38; Text 'Napredne Funkcije'
   Button "Button_1" at 112,438 size 275x137; TextOff 'Rocno Prozenje Branja'
      on Press: function_b14e0dd5("Rocno_Prozenje", 0)
   Button "Button_2" at 493,438 size 275x137; TextOff 'Posodobi Artikel'; Authorization "Visok_Nivo_Autoriteta"
      on Click: ActivateScreen("Lector_Posodobi_Artikel", 0)
   Button "Button_3" at 32,963 size 143x43; TextOff '<<'
      on Press: ActivateScreen("Lector_Branje_Tabela", 0)
   Button "Button_4" at 227,963 size 143x43; TextOff '<< / Glavni Meni'
      on Press: ActivateScreen("Lector_zacetek", 0)
   Button "Button_5" at 879,439 size 275x137; TextOff 'Administracija'
      on Press: ActivateScreen("Lector_Administracija", 0)

screen "Lector_Posodobi_Artikel" 1280x1024, template "Template_LectorStart"
   on GenerateScreen: SetTag("Novi_Artikel_Ime_Artikla_Temp", 0); SetTag("Novi_Artikel_ID_Artikla_Temp", 0); SetTag("Novi_Artikel_Koda_Artikla_Temp", '""')
   TextField "Text field_1" at 504,334 size 253x40; Text 'Posodobi Artikel'
   Button "Button_3" at 32,963 size 143x43; TextOff '<<'
      on Press: ActivateScreen("Lector_Branje_Tabela", 0); function_f23ef4c9()
   Button "Button_4" at 227,963 size 143x43; TextOff '<< / Glavni Meni'
      on Press: ActivateScreen("Lector_zacetek", 0); function_f23ef4c9()
   AlarmView "Alarm view_1" at 330,10 size 600x300
   Button "Button_1" at 556,856 size 178x76; TextOff 'IZBRISI ARTIKEL'; Authorization "Visok_Nivo_Autoriteta"
      on Click: "IZBRISI_Artikel"('Database_ArchiveMessage')
   Button "Button_2" at 556,642 size 178x76; TextOff 'Posodobi'
      on Click: "Posodobi_Artikel"('Database_ArchiveMessage')
   IOField "IO Field" at 313,541 size 284x43; FormatPattern ???????????????????????????????????????????????????????????????????????????????????????????????????????????????????????????????????????????????????????????????????????????????????????????????????????????????????????????????????????????????????????????????
      ProcessValue <- "Novi_Artikel_Ime_Artikla_Temp"
   IOField "IO Field_7" at 60,539 size 219x43; FormatPattern 999
      ProcessValue <- "Novi_Artikel_ID_Artikla_Temp"
      on OnFinishInput: "Posodobi_Iskanje_po_ID"('Database_ArchiveMessage')
   TextField "Text Field_12" at 60,469 size 220x43; Text 'Nr. / No. / ID'
   TextField "Text Field_2" at 313,469 size 284x43; Text 'Nr. / No. / Ime Artikla'
   IOField "IO Field_4" at 630,540 size 580x43; FormatPattern ???????????????????????????????????????????????????????????????????????????????????????????????????????????????????????????????????????????????????????????????????????????????????????????????????????????????????????????????????????????????????????????????
      ProcessValue <- "Novi_Artikel_Koda_Artikla_Temp"
   TextField "Text Field_5" at 630,468 size 580x43; Text 'Nr. / No. / Serijska Stevilka'

screen "Lector_Administracija" 1280x1024, template "Template_LectorStart"
   on GenerateScreen: function_f23ef4c9()
   on ClearScreen: function_f23ef4c9()
   UserView "User view_1" at 22,356 size 1231x508
   Button "Button_1" at 562,890 size 216x70; TextOff 'Odjavi se'
      on Click: function_f23ef4c9()
   Button "Button_3" at 32,963 size 143x43; TextOff '<<'
      on Press: function_efd93a16()
   Button "Button_4" at 227,963 size 143x43; TextOff '<< / Glavni Meni'
      on Press: ActivateScreen("Lector_zacetek", 0)

VB script "S01a_Create_database"
   '////////////////////////////////////////////////////////////////
   ' en: Creating a new database
   ' de: Erstellen einer neuen Datenbank
   ' Created: 19-07-2012
   ' Version: v1.0
   ' Author:  HH
   '////////////////////////////////////////////////////////////////
   
   'Declaration of local tags - Deklarartion von lokalen Variablen
   Dim conn, rst, SQL_Table
   
   On Error Resume Next
   
   Set conn = CreateObject("ADODB.Connection")
   Set rst = CreateObject("ADODB.Recordset")
   
